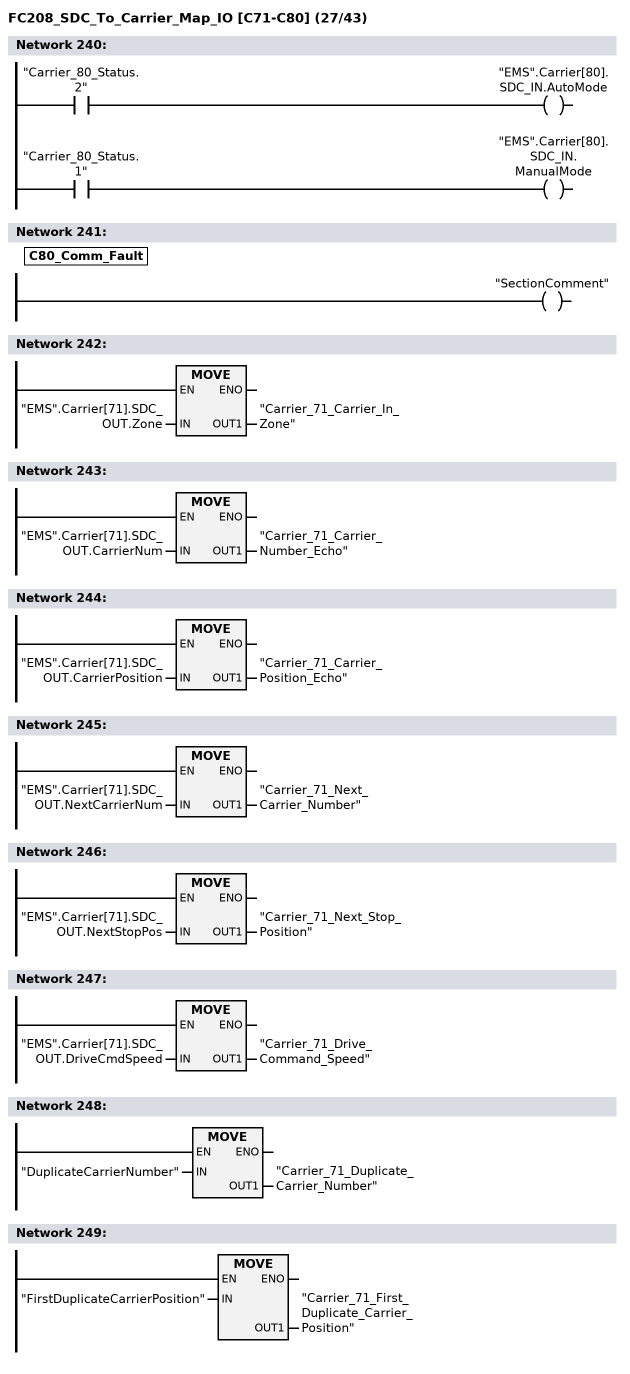
   RUNG wire#powerrail
      Contact( "Carrier_80_Status.2" )
      Coil( "EMS".Carrier[80].SDC_IN.AutoMode )
   END_RUNG
   RUNG wire#powerrail
      Contact( "Carrier_80_Status.1" )
      Coil( "EMS".Carrier[80].SDC_IN.ManualMode )
   END_RUNG
   // the same network as SCL:
   "EMS".Carrier[80].SDC_IN.AutoMode := "Carrier_80_Status.2";
   "EMS".Carrier[80].SDC_IN.ManualMode := "Carrier_80_Status.1";
END_REGION

REGION Network 241
   Label( C80_Comm_Fault )
   RUNG wire#powerrail
      Coil( "SectionComment" )
   END_RUNG
   // the same network as SCL:
   C80_Comm_Fault:
   "SectionComment" := TRUE;
END_REGION

REGION Network 242
   RUNG wire#powerrail
      Move(in := "EMS".Carrier[71].SDC_OUT.Zone, out1 => "Carrier_71_Carrier_In_Zone")
   END_RUNG
   // the same network as SCL:
   "Carrier_71_Carrier_In_Zone" := "EMS".Carrier[71].SDC_OUT.Zone;
END_REGION

REGION Network 243
   RUNG wire#powerrail
      Move(in := "EMS".Carrier[71].SDC_OUT.CarrierNum, out1 => "Carrier_71_Carrier_Number_Echo")
   END_RUNG
   // the same network as SCL:
   "Carrier_71_Carrier_Number_Echo" := "EMS".Carrier[71].SDC_OUT.CarrierNum;
END_REGION

REGION Network 244
   RUNG wire#powerrail
      Move(in := "EMS".Carrier[71].SDC_OUT.CarrierPosition, out1 => "Carrier_71_Carrier_Position_Echo")
   END_RUNG
   // the same network as SCL:
   "Carrier_71_Carrier_Position_Echo" := "EMS".Carrier[71].SDC_OUT.CarrierPosition;
END_REGION

REGION Network 245
   RUNG wire#powerrail
      Move(in := "EMS".Carrier[71].SDC_OUT.NextCarrierNum, out1 => "Carrier_71_Next_Carrier_Number")
   END_RUNG
   // the same network as SCL:
   "Carrier_71_Next_Carrier_Number" := "EMS".Carrier[71].SDC_OUT.NextCarrierNum;
END_REGION

REGION Network 246
   RUNG wire#powerrail
      Move(in := "EMS".Carrier[71].SDC_OUT.NextStopPos, out1 => "Carrier_71_Next_Stop_Position")
   END_RUNG
   // the same network as SCL:
   "Carrier_71_Next_Stop_Position" := "EMS".Carrier[71].SDC_OUT.NextStopPos;
END_REGION

REGION Network 247
   RUNG wire#powerrail
      Move(in := "EMS".Carrier[71].SDC_OUT.DriveCmdSpeed, out1 => "Carrier_71_Drive_Command_Speed")
   END_RUNG
   // the same network as SCL:
   "Carrier_71_Drive_Command_Speed" := "EMS".Carrier[71].SDC_OUT.DriveCmdSpeed;
END_REGION

REGION Network 248
   RUNG wire#powerrail
      Move(in := "DuplicateCarrierNumber", out1 => "Carrier_71_Duplicate_Carrier_Number")
   END_RUNG
   // the same network as SCL:
   "Carrier_71_Duplicate_Carrier_Number" := "DuplicateCarrierNumber";
END_REGION

REGION Network 249
   RUNG wire#powerrail
      Move(in := "FirstDuplicateCarrierPosition", out1 => "Carrier_71_First_Duplicate_Carrier_Position")
   END_RUNG
   // the same network as SCL:
   "Carrier_71_First_Duplicate_Carrier_Position" := "FirstDuplicateCarrierPosition";
END_REGION

REGION Network 250
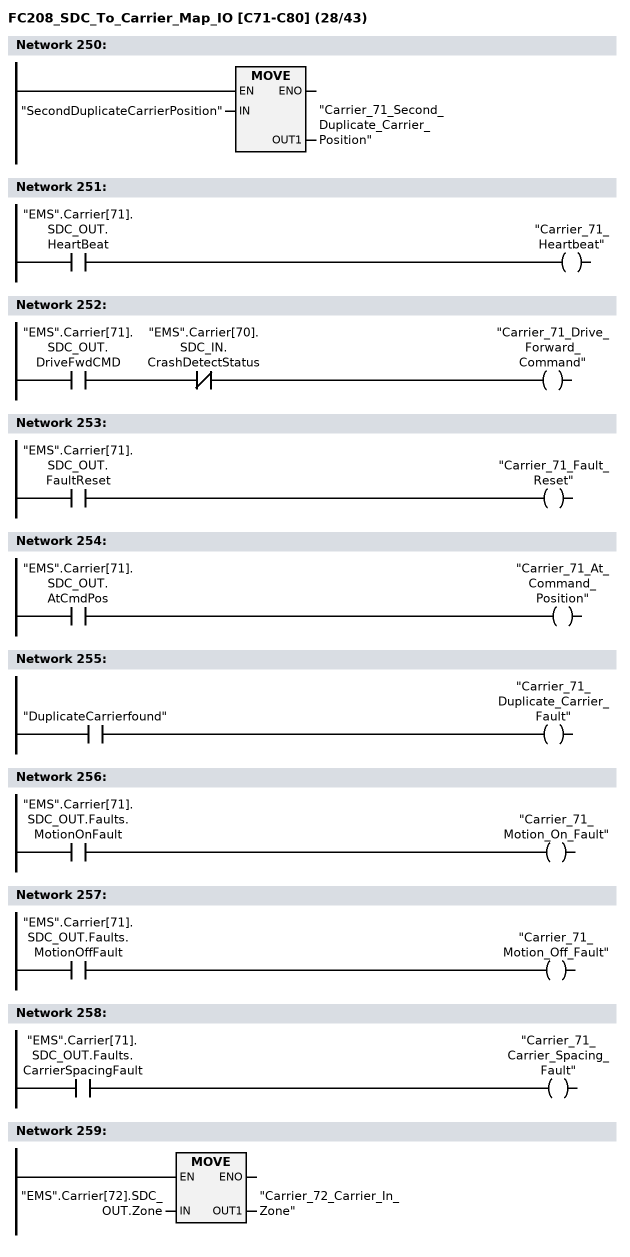
   RUNG wire#powerrail
      Move(in := "SecondDuplicateCarrierPosition", out1 => "Carrier_71_Second_Duplicate_Carrier_Position")
   END_RUNG
   // the same network as SCL:
   "Carrier_71_Second_Duplicate_Carrier_Position" := "SecondDuplicateCarrierPosition";
END_REGION

REGION Network 251
   RUNG wire#powerrail
      Contact( "EMS".Carrier[71].SDC_OUT.HeartBeat )
      Coil( "Carrier_71_Heartbeat" )
   END_RUNG
   // the same network as SCL:
   "Carrier_71_Heartbeat" := "EMS".Carrier[71].SDC_OUT.HeartBeat;
END_REGION

REGION Network 252
   RUNG wire#powerrail
      Contact( "EMS".Carrier[71].SDC_OUT.DriveFwdCMD )
      I_Contact( "EMS".Carrier[70].SDC_IN.CrashDetectStatus )
      Coil( "Carrier_71_Drive_Forward_Command" )
   END_RUNG
   // the same network as SCL:
   "Carrier_71_Drive_Forward_Command" := "EMS".Carrier[71].SDC_OUT.DriveFwdCMD AND NOT "EMS".Carrier[70].SDC_IN.CrashDetectStatus;
END_REGION

REGION Network 253
   RUNG wire#powerrail
      Contact( "EMS".Carrier[71].SDC_OUT.FaultReset )
      Coil( "Carrier_71_Fault_Reset" )
   END_RUNG
   // the same network as SCL:
   "Carrier_71_Fault_Reset" := "EMS".Carrier[71].SDC_OUT.FaultReset;
END_REGION

REGION Network 254
   RUNG wire#powerrail
      Contact( "EMS".Carrier[71].SDC_OUT.AtCmdPos )
      Coil( "Carrier_71_At_Command_Position" )
   END_RUNG
   // the same network as SCL:
   "Carrier_71_At_Command_Position" := "EMS".Carrier[71].SDC_OUT.AtCmdPos;
END_REGION

REGION Network 255
   RUNG wire#powerrail
      Contact( "DuplicateCarrierfound" )
      Coil( "Carrier_71_Duplicate_Carrier_Fault" )
   END_RUNG
   // the same network as SCL:
   "Carrier_71_Duplicate_Carrier_Fault" := "DuplicateCarrierfound";
END_REGION

REGION Network 256
   RUNG wire#powerrail
      Contact( "EMS".Carrier[71].SDC_OUT.Faults.MotionOnFault )
      Coil( "Carrier_71_Motion_On_Fault" )
   END_RUNG
   // the same network as SCL:
   "Carrier_71_Motion_On_Fault" := "EMS".Carrier[71].SDC_OUT.Faults.MotionOnFault;
END_REGION

REGION Network 257
   RUNG wire#powerrail
      Contact( "EMS".Carrier[71].SDC_OUT.Faults.MotionOffFault )
      Coil( "Carrier_71_Motion_Off_Fault" )
   END_RUNG
   // the same network as SCL:
   "Carrier_71_Motion_Off_Fault" := "EMS".Carrier[71].SDC_OUT.Faults.MotionOffFault;
END_REGION

REGION Network 258
   RUNG wire#powerrail
      Contact( "EMS".Carrier[71].SDC_OUT.Faults.CarrierSpacingFault )
      Coil( "Carrier_71_Carrier_Spacing_Fault" )
   END_RUNG
   // the same network as SCL:
   "Carrier_71_Carrier_Spacing_Fault" := "EMS".Carrier[71].SDC_OUT.Faults.CarrierSpacingFault;
END_REGION

REGION Network 259
   RUNG wire#powerrail
      Move(in := "EMS".Carrier[72].SDC_OUT.Zone, out1 => "Carrier_72_Carrier_In_Zone")
   END_RUNG
   // the same network as SCL:
   "Carrier_72_Carrier_In_Zone" := "EMS".Carrier[72].SDC_OUT.Zone;
END_REGION

REGION Network 260
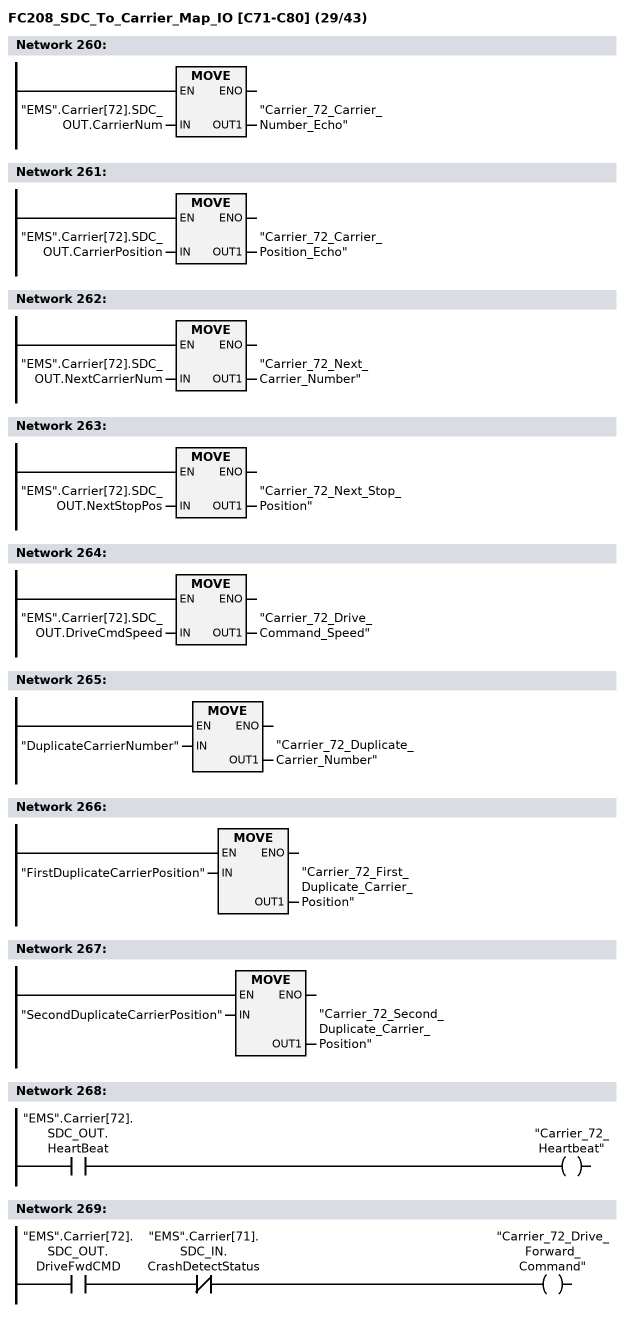
   RUNG wire#powerrail
      Move(in := "EMS".Carrier[72].SDC_OUT.CarrierNum, out1 => "Carrier_72_Carrier_Number_Echo")
   END_RUNG
   // the same network as SCL:
   "Carrier_72_Carrier_Number_Echo" := "EMS".Carrier[72].SDC_OUT.CarrierNum;
END_REGION

REGION Network 261
   RUNG wire#powerrail
      Move(in := "EMS".Carrier[72].SDC_OUT.CarrierPosition, out1 => "Carrier_72_Carrier_Position_Echo")
   END_RUNG
   // the same network as SCL:
   "Carrier_72_Carrier_Position_Echo" := "EMS".Carrier[72].SDC_OUT.CarrierPosition;
END_REGION

REGION Network 262
   RUNG wire#powerrail
      Move(in := "EMS".Carrier[72].SDC_OUT.NextCarrierNum, out1 => "Carrier_72_Next_Carrier_Number")
   END_RUNG
   // the same network as SCL:
   "Carrier_72_Next_Carrier_Number" := "EMS".Carrier[72].SDC_OUT.NextCarrierNum;
END_REGION

REGION Network 263
   RUNG wire#powerrail
      Move(in := "EMS".Carrier[72].SDC_OUT.NextStopPos, out1 => "Carrier_72_Next_Stop_Position")
   END_RUNG
   // the same network as SCL:
   "Carrier_72_Next_Stop_Position" := "EMS".Carrier[72].SDC_OUT.NextStopPos;
END_REGION

REGION Network 264
   RUNG wire#powerrail
      Move(in := "EMS".Carrier[72].SDC_OUT.DriveCmdSpeed, out1 => "Carrier_72_Drive_Command_Speed")
   END_RUNG
   // the same network as SCL:
   "Carrier_72_Drive_Command_Speed" := "EMS".Carrier[72].SDC_OUT.DriveCmdSpeed;
END_REGION

REGION Network 265
   RUNG wire#powerrail
      Move(in := "DuplicateCarrierNumber", out1 => "Carrier_72_Duplicate_Carrier_Number")
   END_RUNG
   // the same network as SCL:
   "Carrier_72_Duplicate_Carrier_Number" := "DuplicateCarrierNumber";
END_REGION

REGION Network 266
   RUNG wire#powerrail
      Move(in := "FirstDuplicateCarrierPosition", out1 => "Carrier_72_First_Duplicate_Carrier_Position")
   END_RUNG
   // the same network as SCL:
   "Carrier_72_First_Duplicate_Carrier_Position" := "FirstDuplicateCarrierPosition";
END_REGION

REGION Network 267
   RUNG wire#powerrail
      Move(in := "SecondDuplicateCarrierPosition", out1 => "Carrier_72_Second_Duplicate_Carrier_Position")
   END_RUNG
   // the same network as SCL:
   "Carrier_72_Second_Duplicate_Carrier_Position" := "SecondDuplicateCarrierPosition";
END_REGION

REGION Network 268
   RUNG wire#powerrail
      Contact( "EMS".Carrier[72].SDC_OUT.HeartBeat )
      Coil( "Carrier_72_Heartbeat" )
   END_RUNG
   // the same network as SCL:
   "Carrier_72_Heartbeat" := "EMS".Carrier[72].SDC_OUT.HeartBeat;
END_REGION

REGION Network 269
   RUNG wire#powerrail
      Contact( "EMS".Carrier[72].SDC_OUT.DriveFwdCMD )
      I_Contact( "EMS".Carrier[71].SDC_IN.CrashDetectStatus )
      Coil( "Carrier_72_Drive_Forward_Command" )
   END_RUNG
   // the same network as SCL:
   "Carrier_72_Drive_Forward_Command" := "EMS".Carrier[72].SDC_OUT.DriveFwdCMD AND NOT "EMS".Carrier[71].SDC_IN.CrashDetectStatus;
END_REGION

REGION Network 270
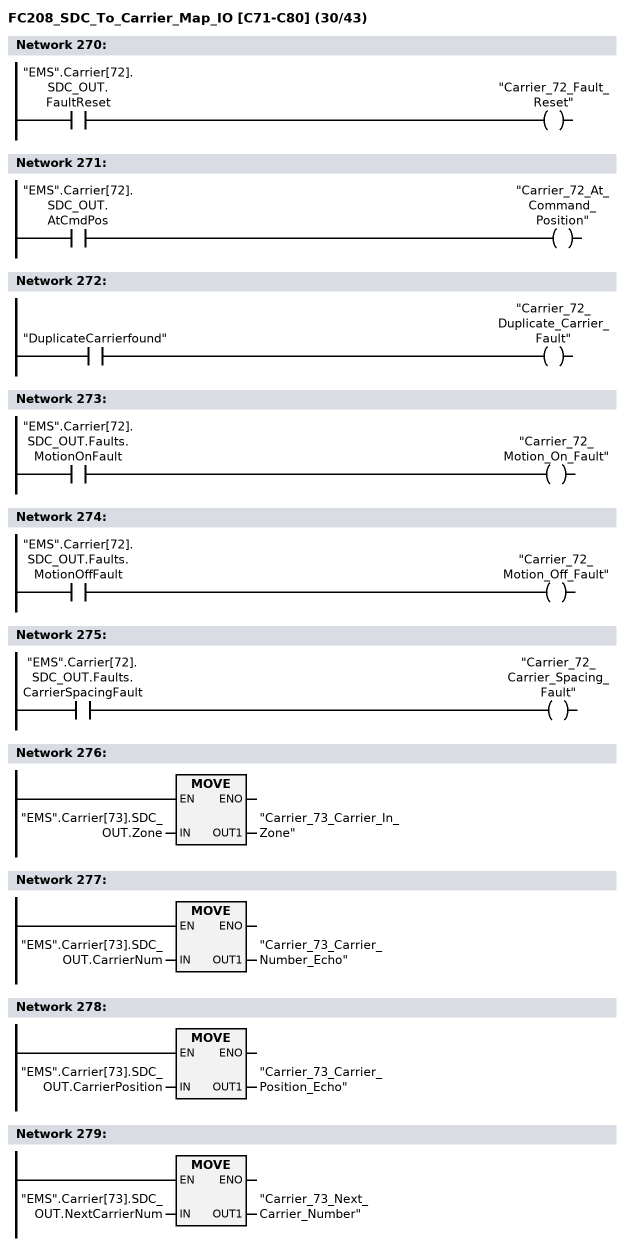
   RUNG wire#powerrail
      Contact( "EMS".Carrier[72].SDC_OUT.FaultReset )
      Coil( "Carrier_72_Fault_Reset" )
   END_RUNG
   // the same network as SCL:
   "Carrier_72_Fault_Reset" := "EMS".Carrier[72].SDC_OUT.FaultReset;
END_REGION

REGION Network 271
   RUNG wire#powerrail
      Contact( "EMS".Carrier[72].SDC_OUT.AtCmdPos )
      Coil( "Carrier_72_At_Command_Position" )
   END_RUNG
   // the same network as SCL:
   "Carrier_72_At_Command_Position" := "EMS".Carrier[72].SDC_OUT.AtCmdPos;
END_REGION

REGION Network 272
   RUNG wire#powerrail
      Contact( "DuplicateCarrierfound" )
      Coil( "Carrier_72_Duplicate_Carrier_Fault" )
   END_RUNG
   // the same network as SCL:
   "Carrier_72_Duplicate_Carrier_Fault" := "DuplicateCarrierfound";
END_REGION

REGION Network 273
   RUNG wire#powerrail
      Contact( "EMS".Carrier[72].SDC_OUT.Faults.MotionOnFault )
      Coil( "Carrier_72_Motion_On_Fault" )
   END_RUNG
   // the same network as SCL:
   "Carrier_72_Motion_On_Fault" := "EMS".Carrier[72].SDC_OUT.Faults.MotionOnFault;
END_REGION

REGION Network 274
   RUNG wire#powerrail
      Contact( "EMS".Carrier[72].SDC_OUT.Faults.MotionOffFault )
      Coil( "Carrier_72_Motion_Off_Fault" )
   END_RUNG
   // the same network as SCL:
   "Carrier_72_Motion_Off_Fault" := "EMS".Carrier[72].SDC_OUT.Faults.MotionOffFault;
END_REGION

REGION Network 275
   RUNG wire#powerrail
      Contact( "EMS".Carrier[72].SDC_OUT.Faults.CarrierSpacingFault )
      Coil( "Carrier_72_Carrier_Spacing_Fault" )
   END_RUNG
   // the same network as SCL:
   "Carrier_72_Carrier_Spacing_Fault" := "EMS".Carrier[72].SDC_OUT.Faults.CarrierSpacingFault;
END_REGION

REGION Network 276
   RUNG wire#powerrail
      Move(in := "EMS".Carrier[73].SDC_OUT.Zone, out1 => "Carrier_73_Carrier_In_Zone")
   END_RUNG
   // the same network as SCL:
   "Carrier_73_Carrier_In_Zone" := "EMS".Carrier[73].SDC_OUT.Zone;
END_REGION

REGION Network 277
   RUNG wire#powerrail
      Move(in := "EMS".Carrier[73].SDC_OUT.CarrierNum, out1 => "Carrier_73_Carrier_Number_Echo")
   END_RUNG
   // the same network as SCL:
   "Carrier_73_Carrier_Number_Echo" := "EMS".Carrier[73].SDC_OUT.CarrierNum;
END_REGION

REGION Network 278
   RUNG wire#powerrail
      Move(in := "EMS".Carrier[73].SDC_OUT.CarrierPosition, out1 => "Carrier_73_Carrier_Position_Echo")
   END_RUNG
   // the same network as SCL:
   "Carrier_73_Carrier_Position_Echo" := "EMS".Carrier[73].SDC_OUT.CarrierPosition;
END_REGION

REGION Network 279
   RUNG wire#powerrail
      Move(in := "EMS".Carrier[73].SDC_OUT.NextCarrierNum, out1 => "Carrier_73_Next_Carrier_Number")
   END_RUNG
   // the same network as SCL:
   "Carrier_73_Next_Carrier_Number" := "EMS".Carrier[73].SDC_OUT.NextCarrierNum;
END_REGION

REGION Network 280
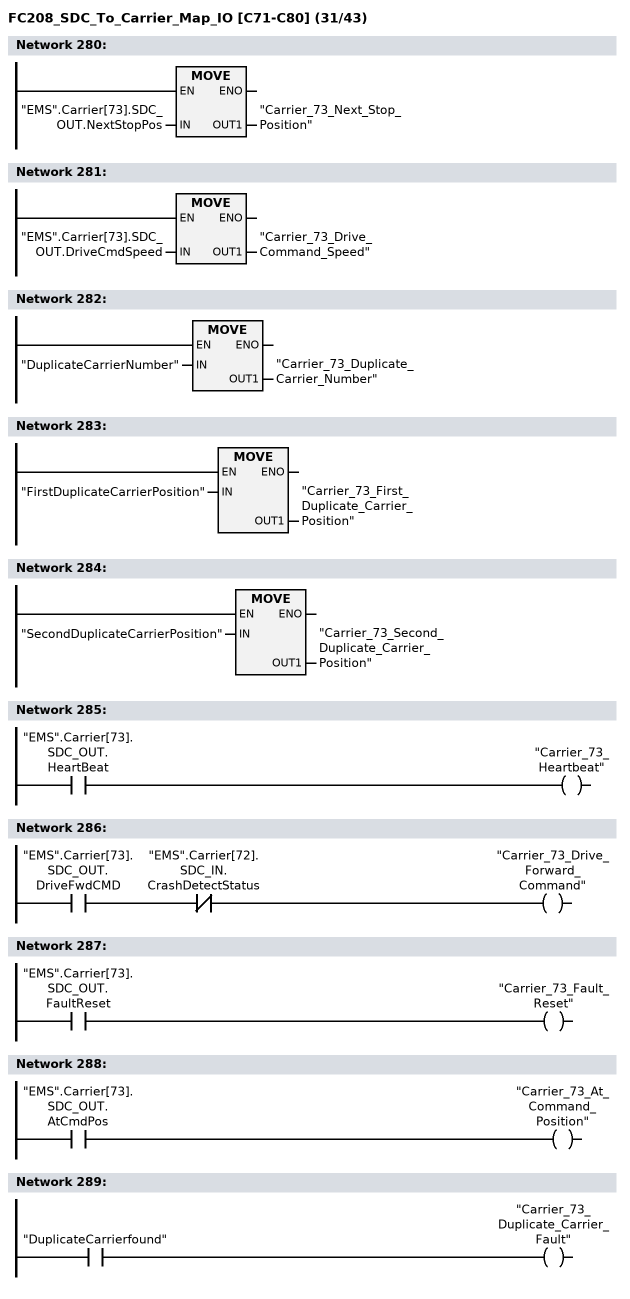
   RUNG wire#powerrail
      Move(in := "EMS".Carrier[73].SDC_OUT.NextStopPos, out1 => "Carrier_73_Next_Stop_Position")
   END_RUNG
   // the same network as SCL:
   "Carrier_73_Next_Stop_Position" := "EMS".Carrier[73].SDC_OUT.NextStopPos;
END_REGION

REGION Network 281
   RUNG wire#powerrail
      Move(in := "EMS".Carrier[73].SDC_OUT.DriveCmdSpeed, out1 => "Carrier_73_Drive_Command_Speed")
   END_RUNG
   // the same network as SCL:
   "Carrier_73_Drive_Command_Speed" := "EMS".Carrier[73].SDC_OUT.DriveCmdSpeed;
END_REGION

REGION Network 282
   RUNG wire#powerrail
      Move(in := "DuplicateCarrierNumber", out1 => "Carrier_73_Duplicate_Carrier_Number")
   END_RUNG
   // the same network as SCL:
   "Carrier_73_Duplicate_Carrier_Number" := "DuplicateCarrierNumber";
END_REGION

REGION Network 283
   RUNG wire#powerrail
      Move(in := "FirstDuplicateCarrierPosition", out1 => "Carrier_73_First_Duplicate_Carrier_Position")
   END_RUNG
   // the same network as SCL:
   "Carrier_73_First_Duplicate_Carrier_Position" := "FirstDuplicateCarrierPosition";
END_REGION

REGION Network 284
   RUNG wire#powerrail
      Move(in := "SecondDuplicateCarrierPosition", out1 => "Carrier_73_Second_Duplicate_Carrier_Position")
   END_RUNG
   // the same network as SCL:
   "Carrier_73_Second_Duplicate_Carrier_Position" := "SecondDuplicateCarrierPosition";
END_REGION

REGION Network 285
   RUNG wire#powerrail
      Contact( "EMS".Carrier[73].SDC_OUT.HeartBeat )
      Coil( "Carrier_73_Heartbeat" )
   END_RUNG
   // the same network as SCL:
   "Carrier_73_Heartbeat" := "EMS".Carrier[73].SDC_OUT.HeartBeat;
END_REGION

REGION Network 286
   RUNG wire#powerrail
      Contact( "EMS".Carrier[73].SDC_OUT.DriveFwdCMD )
      I_Contact( "EMS".Carrier[72].SDC_IN.CrashDetectStatus )
      Coil( "Carrier_73_Drive_Forward_Command" )
   END_RUNG
   // the same network as SCL:
   "Carrier_73_Drive_Forward_Command" := "EMS".Carrier[73].SDC_OUT.DriveFwdCMD AND NOT "EMS".Carrier[72].SDC_IN.CrashDetectStatus;
END_REGION

REGION Network 287
   RUNG wire#powerrail
      Contact( "EMS".Carrier[73].SDC_OUT.FaultReset )
      Coil( "Carrier_73_Fault_Reset" )
   END_RUNG
   // the same network as SCL:
   "Carrier_73_Fault_Reset" := "EMS".Carrier[73].SDC_OUT.FaultReset;
END_REGION

REGION Network 288
   RUNG wire#powerrail
      Contact( "EMS".Carrier[73].SDC_OUT.AtCmdPos )
      Coil( "Carrier_73_At_Command_Position" )
   END_RUNG
   // the same network as SCL:
   "Carrier_73_At_Command_Position" := "EMS".Carrier[73].SDC_OUT.AtCmdPos;
END_REGION

REGION Network 289
   RUNG wire#powerrail
      Contact( "DuplicateCarrierfound" )
      Coil( "Carrier_73_Duplicate_Carrier_Fault" )
   END_RUNG
   // the same network as SCL:
   "Carrier_73_Duplicate_Carrier_Fault" := "DuplicateCarrierfound";
END_REGION

REGION Network 290
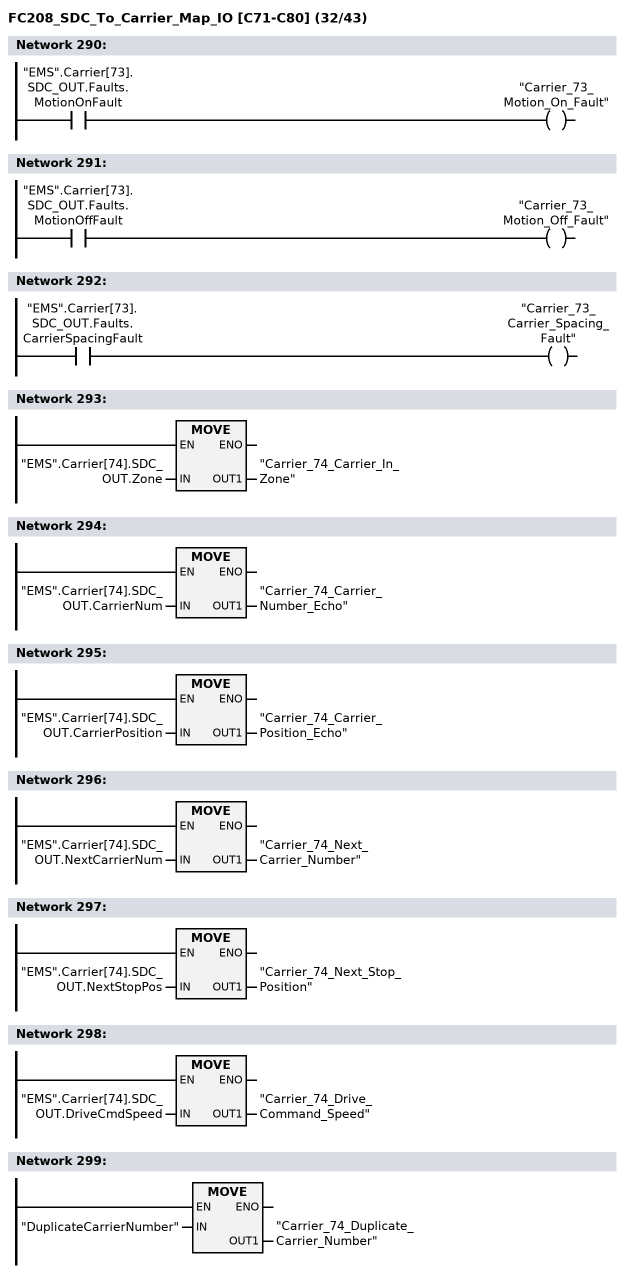
   RUNG wire#powerrail
      Contact( "EMS".Carrier[73].SDC_OUT.Faults.MotionOnFault )
      Coil( "Carrier_73_Motion_On_Fault" )
   END_RUNG
   // the same network as SCL:
   "Carrier_73_Motion_On_Fault" := "EMS".Carrier[73].SDC_OUT.Faults.MotionOnFault;
END_REGION

REGION Network 291
   RUNG wire#powerrail
      Contact( "EMS".Carrier[73].SDC_OUT.Faults.MotionOffFault )
      Coil( "Carrier_73_Motion_Off_Fault" )
   END_RUNG
   // the same network as SCL:
   "Carrier_73_Motion_Off_Fault" := "EMS".Carrier[73].SDC_OUT.Faults.MotionOffFault;
END_REGION

REGION Network 292
   RUNG wire#powerrail
      Contact( "EMS".Carrier[73].SDC_OUT.Faults.CarrierSpacingFault )
      Coil( "Carrier_73_Carrier_Spacing_Fault" )
   END_RUNG
   // the same network as SCL:
   "Carrier_73_Carrier_Spacing_Fault" := "EMS".Carrier[73].SDC_OUT.Faults.CarrierSpacingFault;
END_REGION

REGION Network 293
   RUNG wire#powerrail
      Move(in := "EMS".Carrier[74].SDC_OUT.Zone, out1 => "Carrier_74_Carrier_In_Zone")
   END_RUNG
   // the same network as SCL:
   "Carrier_74_Carrier_In_Zone" := "EMS".Carrier[74].SDC_OUT.Zone;
END_REGION

REGION Network 294
   RUNG wire#powerrail
      Move(in := "EMS".Carrier[74].SDC_OUT.CarrierNum, out1 => "Carrier_74_Carrier_Number_Echo")
   END_RUNG
   // the same network as SCL:
   "Carrier_74_Carrier_Number_Echo" := "EMS".Carrier[74].SDC_OUT.CarrierNum;
END_REGION

REGION Network 295
   RUNG wire#powerrail
      Move(in := "EMS".Carrier[74].SDC_OUT.CarrierPosition, out1 => "Carrier_74_Carrier_Position_Echo")
   END_RUNG
   // the same network as SCL:
   "Carrier_74_Carrier_Position_Echo" := "EMS".Carrier[74].SDC_OUT.CarrierPosition;
END_REGION

REGION Network 296
   RUNG wire#powerrail
      Move(in := "EMS".Carrier[74].SDC_OUT.NextCarrierNum, out1 => "Carrier_74_Next_Carrier_Number")
   END_RUNG
   // the same network as SCL:
   "Carrier_74_Next_Carrier_Number" := "EMS".Carrier[74].SDC_OUT.NextCarrierNum;
END_REGION

REGION Network 297
   RUNG wire#powerrail
      Move(in := "EMS".Carrier[74].SDC_OUT.NextStopPos, out1 => "Carrier_74_Next_Stop_Position")
   END_RUNG
   // the same network as SCL:
   "Carrier_74_Next_Stop_Position" := "EMS".Carrier[74].SDC_OUT.NextStopPos;
END_REGION

REGION Network 298
   RUNG wire#powerrail
      Move(in := "EMS".Carrier[74].SDC_OUT.DriveCmdSpeed, out1 => "Carrier_74_Drive_Command_Speed")
   END_RUNG
   // the same network as SCL:
   "Carrier_74_Drive_Command_Speed" := "EMS".Carrier[74].SDC_OUT.DriveCmdSpeed;
END_REGION

REGION Network 299
   RUNG wire#powerrail
      Move(in := "DuplicateCarrierNumber", out1 => "Carrier_74_Duplicate_Carrier_Number")
   END_RUNG
   // the same network as SCL:
   "Carrier_74_Duplicate_Carrier_Number" := "DuplicateCarrierNumber";
END_REGION

REGION Network 300
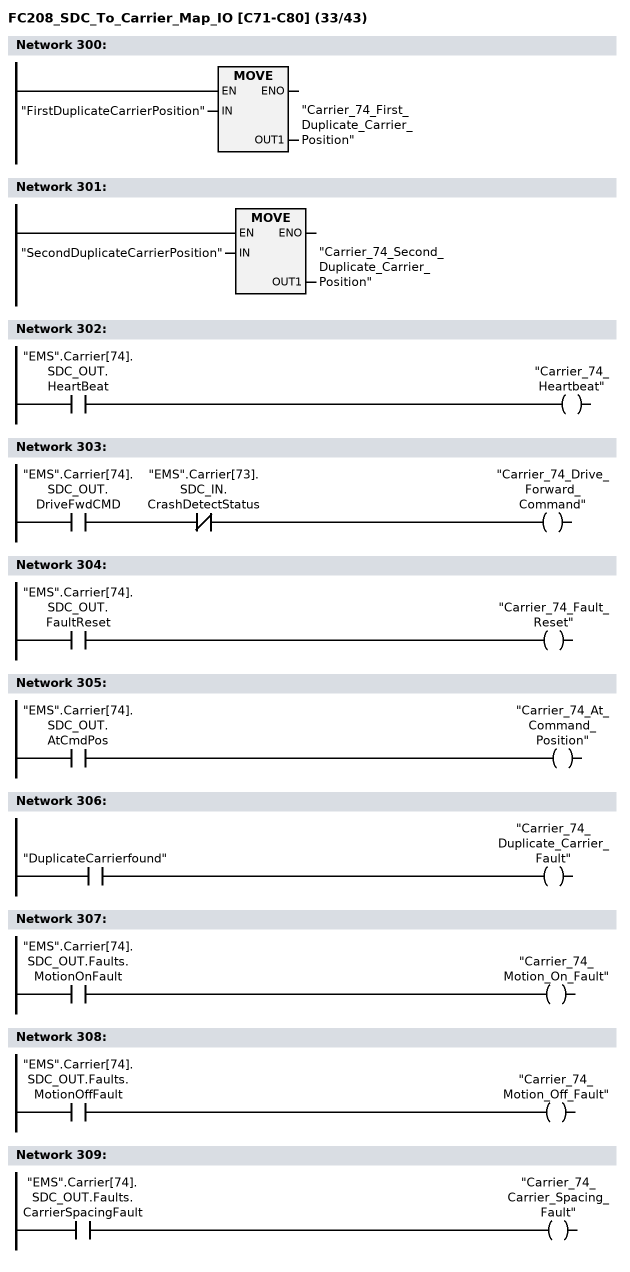
   RUNG wire#powerrail
      Move(in := "FirstDuplicateCarrierPosition", out1 => "Carrier_74_First_Duplicate_Carrier_Position")
   END_RUNG
   // the same network as SCL:
   "Carrier_74_First_Duplicate_Carrier_Position" := "FirstDuplicateCarrierPosition";
END_REGION

REGION Network 301
   RUNG wire#powerrail
      Move(in := "SecondDuplicateCarrierPosition", out1 => "Carrier_74_Second_Duplicate_Carrier_Position")
   END_RUNG
   // the same network as SCL:
   "Carrier_74_Second_Duplicate_Carrier_Position" := "SecondDuplicateCarrierPosition";
END_REGION

REGION Network 302
   RUNG wire#powerrail
      Contact( "EMS".Carrier[74].SDC_OUT.HeartBeat )
      Coil( "Carrier_74_Heartbeat" )
   END_RUNG
   // the same network as SCL:
   "Carrier_74_Heartbeat" := "EMS".Carrier[74].SDC_OUT.HeartBeat;
END_REGION

REGION Network 303
   RUNG wire#powerrail
      Contact( "EMS".Carrier[74].SDC_OUT.DriveFwdCMD )
      I_Contact( "EMS".Carrier[73].SDC_IN.CrashDetectStatus )
      Coil( "Carrier_74_Drive_Forward_Command" )
   END_RUNG
   // the same network as SCL:
   "Carrier_74_Drive_Forward_Command" := "EMS".Carrier[74].SDC_OUT.DriveFwdCMD AND NOT "EMS".Carrier[73].SDC_IN.CrashDetectStatus;
END_REGION

REGION Network 304
   RUNG wire#powerrail
      Contact( "EMS".Carrier[74].SDC_OUT.FaultReset )
      Coil( "Carrier_74_Fault_Reset" )
   END_RUNG
   // the same network as SCL:
   "Carrier_74_Fault_Reset" := "EMS".Carrier[74].SDC_OUT.FaultReset;
END_REGION

REGION Network 305
   RUNG wire#powerrail
      Contact( "EMS".Carrier[74].SDC_OUT.AtCmdPos )
      Coil( "Carrier_74_At_Command_Position" )
   END_RUNG
   // the same network as SCL:
   "Carrier_74_At_Command_Position" := "EMS".Carrier[74].SDC_OUT.AtCmdPos;
END_REGION

REGION Network 306
   RUNG wire#powerrail
      Contact( "DuplicateCarrierfound" )
      Coil( "Carrier_74_Duplicate_Carrier_Fault" )
   END_RUNG
   // the same network as SCL:
   "Carrier_74_Duplicate_Carrier_Fault" := "DuplicateCarrierfound";
END_REGION

REGION Network 307
   RUNG wire#powerrail
      Contact( "EMS".Carrier[74].SDC_OUT.Faults.MotionOnFault )
      Coil( "Carrier_74_Motion_On_Fault" )
   END_RUNG
   // the same network as SCL:
   "Carrier_74_Motion_On_Fault" := "EMS".Carrier[74].SDC_OUT.Faults.MotionOnFault;
END_REGION

REGION Network 308
   RUNG wire#powerrail
      Contact( "EMS".Carrier[74].SDC_OUT.Faults.MotionOffFault )
      Coil( "Carrier_74_Motion_Off_Fault" )
   END_RUNG
   // the same network as SCL:
   "Carrier_74_Motion_Off_Fault" := "EMS".Carrier[74].SDC_OUT.Faults.MotionOffFault;
END_REGION

REGION Network 309
   RUNG wire#powerrail
      Contact( "EMS".Carrier[74].SDC_OUT.Faults.CarrierSpacingFault )
      Coil( "Carrier_74_Carrier_Spacing_Fault" )
   END_RUNG
   // the same network as SCL:
   "Carrier_74_Carrier_Spacing_Fault" := "EMS".Carrier[74].SDC_OUT.Faults.CarrierSpacingFault;
END_REGION

REGION Network 310
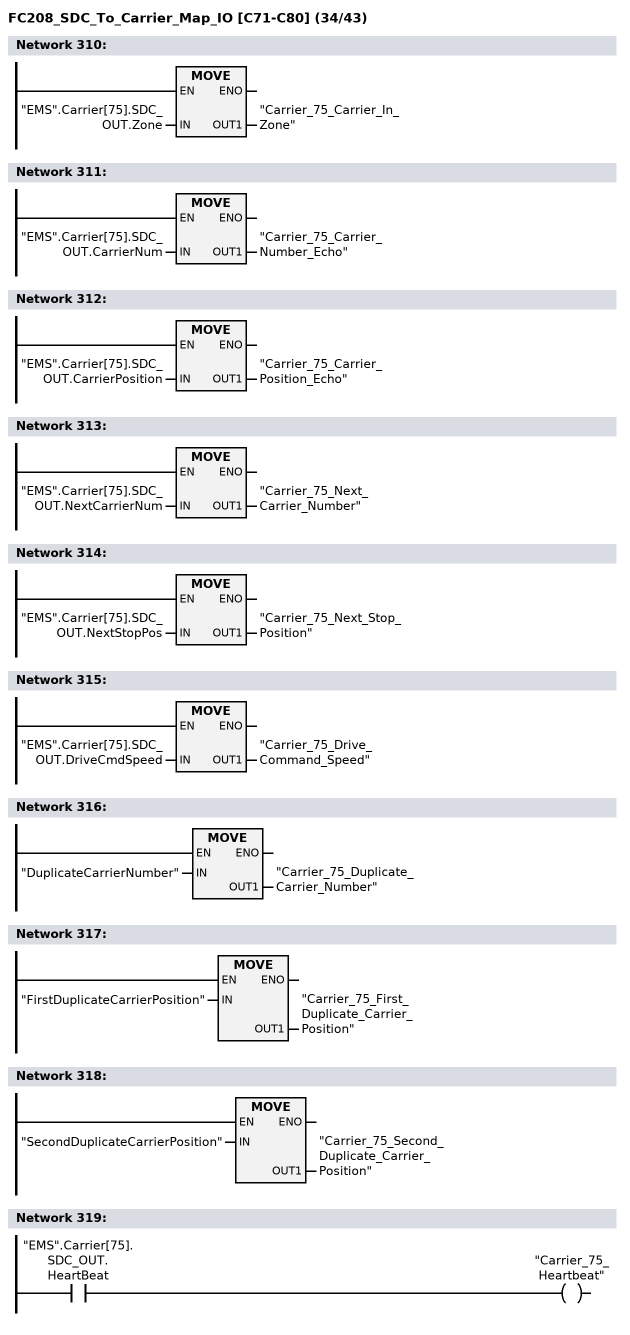
   RUNG wire#powerrail
      Move(in := "EMS".Carrier[75].SDC_OUT.Zone, out1 => "Carrier_75_Carrier_In_Zone")
   END_RUNG
   // the same network as SCL:
   "Carrier_75_Carrier_In_Zone" := "EMS".Carrier[75].SDC_OUT.Zone;
END_REGION

REGION Network 311
   RUNG wire#powerrail
      Move(in := "EMS".Carrier[75].SDC_OUT.CarrierNum, out1 => "Carrier_75_Carrier_Number_Echo")
   END_RUNG
   // the same network as SCL:
   "Carrier_75_Carrier_Number_Echo" := "EMS".Carrier[75].SDC_OUT.CarrierNum;
END_REGION

REGION Network 312
   RUNG wire#powerrail
      Move(in := "EMS".Carrier[75].SDC_OUT.CarrierPosition, out1 => "Carrier_75_Carrier_Position_Echo")
   END_RUNG
   // the same network as SCL:
   "Carrier_75_Carrier_Position_Echo" := "EMS".Carrier[75].SDC_OUT.CarrierPosition;
END_REGION

REGION Network 313
   RUNG wire#powerrail
      Move(in := "EMS".Carrier[75].SDC_OUT.NextCarrierNum, out1 => "Carrier_75_Next_Carrier_Number")
   END_RUNG
   // the same network as SCL:
   "Carrier_75_Next_Carrier_Number" := "EMS".Carrier[75].SDC_OUT.NextCarrierNum;
END_REGION

REGION Network 314
   RUNG wire#powerrail
      Move(in := "EMS".Carrier[75].SDC_OUT.NextStopPos, out1 => "Carrier_75_Next_Stop_Position")
   END_RUNG
   // the same network as SCL:
   "Carrier_75_Next_Stop_Position" := "EMS".Carrier[75].SDC_OUT.NextStopPos;
END_REGION

REGION Network 315
   RUNG wire#powerrail
      Move(in := "EMS".Carrier[75].SDC_OUT.DriveCmdSpeed, out1 => "Carrier_75_Drive_Command_Speed")
   END_RUNG
   // the same network as SCL:
   "Carrier_75_Drive_Command_Speed" := "EMS".Carrier[75].SDC_OUT.DriveCmdSpeed;
END_REGION

REGION Network 316
   RUNG wire#powerrail
      Move(in := "DuplicateCarrierNumber", out1 => "Carrier_75_Duplicate_Carrier_Number")
   END_RUNG
   // the same network as SCL:
   "Carrier_75_Duplicate_Carrier_Number" := "DuplicateCarrierNumber";
END_REGION

REGION Network 317
   RUNG wire#powerrail
      Move(in := "FirstDuplicateCarrierPosition", out1 => "Carrier_75_First_Duplicate_Carrier_Position")
   END_RUNG
   // the same network as SCL:
   "Carrier_75_First_Duplicate_Carrier_Position" := "FirstDuplicateCarrierPosition";
END_REGION

REGION Network 318
   RUNG wire#powerrail
      Move(in := "SecondDuplicateCarrierPosition", out1 => "Carrier_75_Second_Duplicate_Carrier_Position")
   END_RUNG
   // the same network as SCL:
   "Carrier_75_Second_Duplicate_Carrier_Position" := "SecondDuplicateCarrierPosition";
END_REGION

REGION Network 319
   RUNG wire#powerrail
      Contact( "EMS".Carrier[75].SDC_OUT.HeartBeat )
      Coil( "Carrier_75_Heartbeat" )
   END_RUNG
   // the same network as SCL:
   "Carrier_75_Heartbeat" := "EMS".Carrier[75].SDC_OUT.HeartBeat;
END_REGION

REGION Network 320
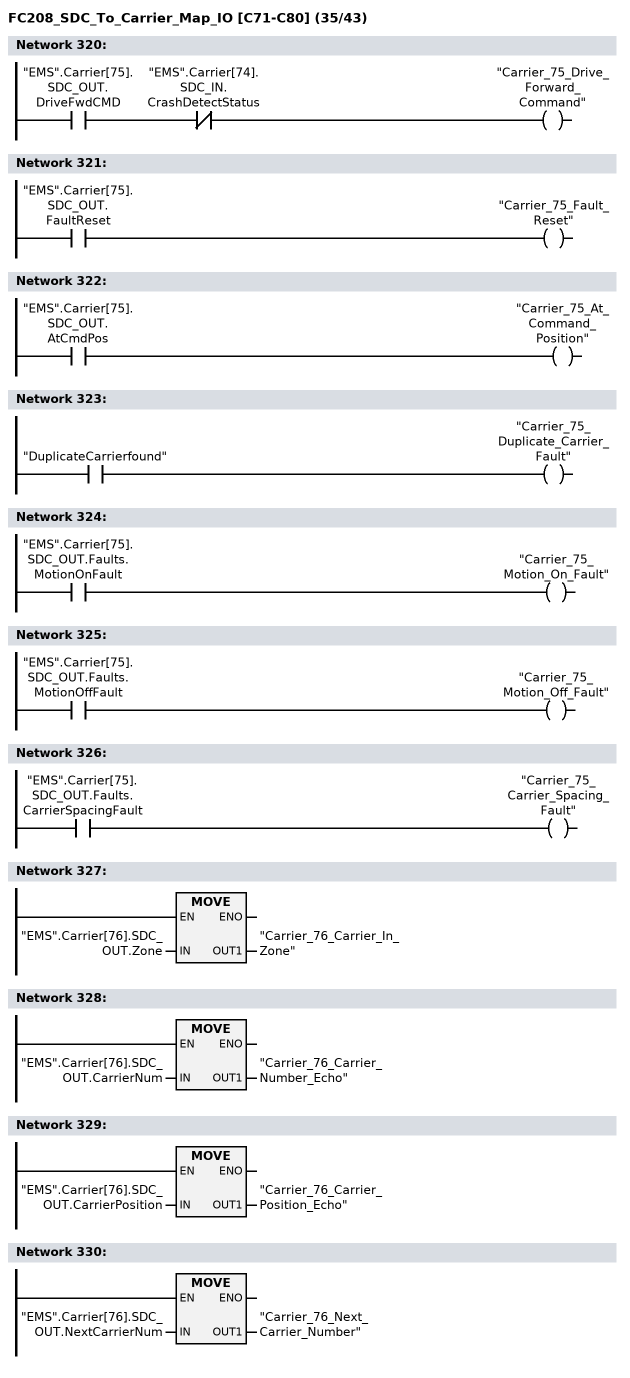
   RUNG wire#powerrail
      Contact( "EMS".Carrier[75].SDC_OUT.DriveFwdCMD )
      I_Contact( "EMS".Carrier[74].SDC_IN.CrashDetectStatus )
      Coil( "Carrier_75_Drive_Forward_Command" )
   END_RUNG
   // the same network as SCL:
   "Carrier_75_Drive_Forward_Command" := "EMS".Carrier[75].SDC_OUT.DriveFwdCMD AND NOT "EMS".Carrier[74].SDC_IN.CrashDetectStatus;
END_REGION

REGION Network 321
   RUNG wire#powerrail
      Contact( "EMS".Carrier[75].SDC_OUT.FaultReset )
      Coil( "Carrier_75_Fault_Reset" )
   END_RUNG
   // the same network as SCL:
   "Carrier_75_Fault_Reset" := "EMS".Carrier[75].SDC_OUT.FaultReset;
END_REGION

REGION Network 322
   RUNG wire#powerrail
      Contact( "EMS".Carrier[75].SDC_OUT.AtCmdPos )
      Coil( "Carrier_75_At_Command_Position" )
   END_RUNG
   // the same network as SCL:
   "Carrier_75_At_Command_Position" := "EMS".Carrier[75].SDC_OUT.AtCmdPos;
END_REGION

REGION Network 323
   RUNG wire#powerrail
      Contact( "DuplicateCarrierfound" )
      Coil( "Carrier_75_Duplicate_Carrier_Fault" )
   END_RUNG
   // the same network as SCL:
   "Carrier_75_Duplicate_Carrier_Fault" := "DuplicateCarrierfound";
END_REGION

REGION Network 324
   RUNG wire#powerrail
      Contact( "EMS".Carrier[75].SDC_OUT.Faults.MotionOnFault )
      Coil( "Carrier_75_Motion_On_Fault" )
   END_RUNG
   // the same network as SCL:
   "Carrier_75_Motion_On_Fault" := "EMS".Carrier[75].SDC_OUT.Faults.MotionOnFault;
END_REGION

REGION Network 325
   RUNG wire#powerrail
      Contact( "EMS".Carrier[75].SDC_OUT.Faults.MotionOffFault )
      Coil( "Carrier_75_Motion_Off_Fault" )
   END_RUNG
   // the same network as SCL:
   "Carrier_75_Motion_Off_Fault" := "EMS".Carrier[75].SDC_OUT.Faults.MotionOffFault;
END_REGION

REGION Network 326
   RUNG wire#powerrail
      Contact( "EMS".Carrier[75].SDC_OUT.Faults.CarrierSpacingFault )
      Coil( "Carrier_75_Carrier_Spacing_Fault" )
   END_RUNG
   // the same network as SCL:
   "Carrier_75_Carrier_Spacing_Fault" := "EMS".Carrier[75].SDC_OUT.Faults.CarrierSpacingFault;
END_REGION

REGION Network 327
   RUNG wire#powerrail
      Move(in := "EMS".Carrier[76].SDC_OUT.Zone, out1 => "Carrier_76_Carrier_In_Zone")
   END_RUNG
   // the same network as SCL:
   "Carrier_76_Carrier_In_Zone" := "EMS".Carrier[76].SDC_OUT.Zone;
END_REGION

REGION Network 328
   RUNG wire#powerrail
      Move(in := "EMS".Carrier[76].SDC_OUT.CarrierNum, out1 => "Carrier_76_Carrier_Number_Echo")
   END_RUNG
   // the same network as SCL:
   "Carrier_76_Carrier_Number_Echo" := "EMS".Carrier[76].SDC_OUT.CarrierNum;
END_REGION

REGION Network 329
   RUNG wire#powerrail
      Move(in := "EMS".Carrier[76].SDC_OUT.CarrierPosition, out1 => "Carrier_76_Carrier_Position_Echo")
   END_RUNG
   // the same network as SCL:
   "Carrier_76_Carrier_Position_Echo" := "EMS".Carrier[76].SDC_OUT.CarrierPosition;
END_REGION

REGION Network 330
   RUNG wire#powerrail
      Move(in := "EMS".Carrier[76].SDC_OUT.NextCarrierNum, out1 => "Carrier_76_Next_Carrier_Number")
   END_RUNG
   // the same network as SCL:
   "Carrier_76_Next_Carrier_Number" := "EMS".Carrier[76].SDC_OUT.NextCarrierNum;
END_REGION

REGION Network 331
